           #temp_text2 := #Cfg_MessagePrefix.MessagePrefix[#temp_Language];
           IF LEN(#temp_text2) = 0 THEN #temp_text2 := ' ';  END_IF;

           #temp_text3 := #Cfg_Event.Message[#temp_Language];
           IF LEN(#temp_text3) = 0 THEN #temp_text3 := ' ';  END_IF;

        #In_EventStatus.Sts_Events[#Event_Number].Message := CONCAT(IN1 := #temp_text1, IN2 := #temp_text2, IN3 := #temp_text3);   // CONCAT (Cfg_MessagePrefix, Cfg_Event.Message);    
        //  #In_EventStatus.Sts_Events[#Event_Number].Message := CONCAT(IN1 := #temp_text1, IN2 := #Cfg_MessagePrefix.Language[#temp_Language], IN3 := #Cfg_Event.Message[#temp_Language]);   // CONCAT (Cfg_MessagePrefix, Cfg_Event.Message); 

           #In_EventStatus.Sts_Events[#Event_Number].Trigger := TRUE;                      // Set trigger to 1 
           #In_EventStatus.Sts_Events[#Event_Number].DateTime := #Event_CurDateTime;         // Update with the current time
           #In_EventStatus.Sts_Events[#Event_Number].AckDateTime := DT#1990-1-1-0:0:0.0;       // clear the acknowledge time value 
           END_IF;

      #Sts_Active   := TRUE;                            // set the status active bit
      #Sts_Latched  := TRUE;                            // set the status latched bit
      #In_EventStatus.Wrk_UpdateEventListID := #In_EventStatus.Wrk_UpdateEventListID+1;  // increment the work update listID


       CASE DINT_TO_INT(#Cfg_Event.Category) OF                     // set the appropriate category lateched bit 
           0: #In_EventStatus.Sts_Category_0_Latched :=1;
           1: #In_EventStatus.Sts_Category_1_Latched :=1;
           2: #In_EventStatus.Sts_Category_2_Latched :=1;
           3: #In_EventStatus.Sts_Category_3_Latched :=1;
           4: #In_EventStatus.Sts_Category_4_Latched :=1;
           5: #In_EventStatus.Sts_Category_5_Latched :=1;
           6: #In_EventStatus.Sts_Category_6_Latched :=1;
           7: #In_EventStatus.Sts_Category_7_Latched :=1;
           8: #In_EventStatus.Sts_Category_8_Latched :=1;
           9: #In_EventStatus.Sts_Category_9_Latched :=1;
       END_CASE;
   END_IF;                            // End "IF NOT (Sts_Active)"


   END_IF;                             // End "IF NOT(EnableIn) "


   //----------------------------------------------------- 
   ENO:= true;          // Set the ENO output
END_FUNCTION_BLOCK

FUNCTION_BLOCK "FB_TR88_CPG_EventManager"   // FB3102, SCL
TITLE = PackML EventManager (TR88 CPG Template)
{ S7_Optimized_Access := 'TRUE' }
AUTHOR : FoodBev
FAMILY : ISATR88e
NAME : EventMgr
VERSION : 1.81
// Takes the event information from the control modules (from FB_Event) and will create one list of events for the equipment module. It summarizes the data by finding the equipment module first out event and summarizes which category of events are active. This FB will also send reset commands to unlatch the control module events. Only one instance of this FB should be programmed per equipment module for each event type, for example one for alarms, one for warnings, etc.
   VAR_INPUT
      Cmd_Reset : Bool;   // Reset Command
      Cmd_ClearFirstOutEvents : Bool;   // Command to clear First Out events
      FirstScanBit : Bool;   // Bit used to tell logic that this is the firt scan of PLC
      Cfg_MessagePrefix : "UDT_TR88_CPG_Message_Prefix";   // Message Prefix value for event messages multi-lingual
      Cfg_Language : Int;   // Current Langage: 0=EN, 1=SP/ES, 2=DE, 3=FR, 4=IT
   END_VAR
   VAR_OUTPUT
      Sts_Category_0_Latched : Bool;   // Event Category Status (on until reset cmd) - CAT 0
      Sts_Category_1_Latched : Bool;   // Event Category Status (on until reset cmd) - CAT 1
      Sts_Category_2_Latched : Bool;   // Event Category Status (on until reset cmd) - CAT 2
      Sts_Category_3_Latched : Bool;   // Event Category Status (on until reset cmd) - CAT 3
      Sts_Category_4_Latched : Bool;   // Event Category Status (on until reset cmd) - CAT 4
      Sts_Category_5_Latched : Bool;   // Event Category Status (on until reset cmd) - CAT 5
      Sts_Category_6_Latched : Bool;   // Event Category Status (on until reset cmd) - CAT 6
      Sts_Category_7_Latched : Bool;   // Event Category Status (on until reset cmd) - CAT 7
      Sts_Category_8_Latched : Bool;   // Event Category Status (on until reset cmd) - CAT 8
      Sts_Category_9_Latched : Bool;   // Event Category Status (on until reset cmd) - CAT 9
      Sts_Category_0_NotLatched : Bool;   // Event Cat Status, not latched (=active event status) - CAT 0
      Sts_Category_1_NotLatched : Bool;   // Event Cat Status, not latched (=active event status) - CAT 1
      Sts_Category_2_NotLatched : Bool;   // Event Cat Status, not latched (=active event status) - CAT 2
      Sts_Category_3_NotLatched : Bool;   // Event Cat Status, not latched (=active event status) - CAT 3
      Sts_Category_4_NotLatched : Bool;   // Event Cat Status, not latched (=active event status) - CAT 4
      Sts_Category_5_NotLatched : Bool;   // Event Cat Status, not latched (=active event status) - CAT 5
      Sts_Category_6_NotLatched : Bool;   // Event Cat Status, not latched (=active event status) - CAT 6
      Sts_Category_7_NotLatched : Bool;   // Event Cat Status, not latched (=active event status) - CAT 7
      Sts_Category_8_NotLatched : Bool;   // Event Cat Status, not latched (=active event status) - CAT 8
      Sts_Category_9_NotLatched : Bool;   // Event Cat Status, not latched (=active event status) - CAT 9
      Sts_NumEvents : Int;   // Number of event in the In_EventStatus list
      Sts_CurrentActiveEvent : Bool;   // Status - TRUE = if any active events
      Sts_error : Bool;   // FB Error exist
      Sts_errorCode : DInt;   // FB Error code
   END_VAR
   VAR_IN_OUT
      In_EventStatus : "UDT_TR88_CPG_EventStatus";   // Working event list data section
   END_VAR
   VAR
      EventCategory : Int;
      Index_AllEvents : Int;
      Index_ClearActiveEvents : Int;
      Index_ClearFirstOut : Int;
      NumEvents : Int;   // Max # of Events
      Prev_CmdReset : Bool;
      Prev_NumEvents : Int;
      Prev_UpdateEventListID : Int;
      UpdateEventList : Bool;
      ZeroEvent : "UDT_TR88_CPG_Event";   // Null Event
   END_VAR
   VAR_TEMP
      "step" : Int;
      temp_text1 : String[30];
      temp_text2 : String[30];
      tempAnyPointer : DInt;   // temp Any poninter for FC_Array_Length call.
   END_VAR
BEGIN
   // ============================================================================ 
   // FUNCTION_BLOCK "FB_PMLe_EventManager"  
   // ---------------------------------------------------------------------------
   // Siemens Industry, Inc.
   // Food & Beverage VSS
   // ---------------------------------------------------------------------------
   // FUNCTIONALITY:  
   // Function Block to control EventManager function.
   // ---------------------------------------------------------------------------
   // change log table:
   // version        date          expert in charge        changes applied
   //  1.7         2012-08-22          M.Pieper           Matches Rev 1.7
   //                                                     Added Multi-Lingual support
   //  1.8       2013.07.31            M.Pieper           Removed EM message prefix logic
   //  1.81      2015-01-27            M.Pieper           Updated S7-1500 Array Size Logic.
   // ===========================================================================
   (*
   THIS SOFTWARE IS PROVIDED "AS IS" AND WITHOUT WARRANTIES OF ANY KIND, WHETHER EXPRESS OR IMPLIED.

   General information -
       Note :  the standard applications are NOT binding AND DO NOT claim TO be complete regarding configuration, equipment OR any eventuality which may arise. 
       The standard applications DO NOT represent specific customer solutions, but are only intended TO provide support FOR typical tasks. You are responsible 
       FOR the proper operation OF the described products. These standard applications DO NOT relieve you OF your responsibility regarding the safe handling 
       when using, installing operating AND maintaining the equipment. BY using these standard applications, you agree that Siemens cannot be made liable FOR 
       possible damage beyond the mentioned liability clause. We reserve the right TO make changes AND revisions TO these standard applications at Any Time 
       without prior notice. In the CASE OF Any differences between the suggestions made in these standard applications AND other publications from Siemens, 
       such as catalogs, the contents OF the other documentation have priority.

   Warranty conditions, liability, AND support -
      IF the application has been made available free OF charge, the following applies:
      * We DO NOT provide a warranty FOR Any OF the information contained in this document.
      * All other rights AND claims against Siemens AG irrespective OF legal basis are excluded. In particular claims FOR damages against Siemens AG 
      in the CASE OF Product outage, downtime, loss OF profit, either directly, indirectly OR consequential damage are excluded.
      * This does NOT apply when liability is compulsory BY law, e. g. in the CASE OF the Product liability act, premeditation, an act OF gross negligence 
      BY superiors AND managerial staff OF Siemens AG OR in cases OF fraudulent concealment OF defects.
      * This limitation OF liability also applies TO sub-contractors, suppliers, delegates, superiors AND managerial staff OF Siemens AG.
      German law shall apply TO this agreement FOR customers with head offices in Germany; Swiss law FOR customers with head offices outside Germany. 
      Application OF the United Nations Convention on Contracts FOR the International Sale OF Goods as OF 11.04.1980 (CISG) is excluded.
   *)

   // ===========================================================================
   //  Begin the LOGIC section:
   // First Scan Logic Logic (only ran on 1st scan of PLC)
   IF #FirstScanBit THEN                   //  First Scan bit set?
       #In_EventStatus.Wrk_ResetID := #In_EventStatus.Wrk_ResetID + 1;            // increment the Work Reset ID
       #In_EventStatus.Wrk_UpdateEventListID := #In_EventStatus.Wrk_UpdateEventListID + 1; // increment the Work UpdateList ID
       #In_EventStatus.Sts_NumAllEvents := 0;                                        // Reset the number of all events value
       // Determine the Number of Sts_Events for given alarm/warning area
       // S7-1500 Code: 
       "FC_ArrayLength_S7-1500"(Array_ToBe_Sized := #In_EventStatus.Sts_Events,
                                ArraySize => #In_EventStatus.Wrk_EventArraySize);
       RETURN;                            // Exit the FB call
   END_IF;                              // End the first scan section


   //---------------------------------------------------------------------------------
   // Main Logic Section

   // Update the message prefix for the current language
   #In_EventStatus.Wrk_LanguageSelection := #Cfg_Language;
   #In_EventStatus.Wrk_MessagePrefix := #Cfg_MessagePrefix.MessagePrefix[#In_EventStatus.Wrk_LanguageSelection];

   // Upon a reset command, reset the latched status bits and clear the event list
   IF #Cmd_Reset THEN
       #In_EventStatus.Sts_Category_0_Latched := 0;
       #In_EventStatus.Sts_Category_1_Latched := 0;
       #In_EventStatus.Sts_Category_2_Latched := 0;
       #In_EventStatus.Sts_Category_3_Latched := 0;
       #In_EventStatus.Sts_Category_4_Latched := 0;
       #In_EventStatus.Sts_Category_5_Latched := 0;
       #In_EventStatus.Sts_Category_6_Latched := 0;
       #In_EventStatus.Sts_Category_7_Latched := 0;
       #In_EventStatus.Sts_Category_8_Latched := 0;
       #In_EventStatus.Sts_Category_9_Latched := 0;

       IF NOT (#Prev_CmdReset) THEN                             // Clear the zero event
           #In_EventStatus.Out_ZeroEvent := #ZeroEvent;
           // String seperation variable not added.
       END_IF;
   END_IF;                      // End IF Cmd_Reset.... 


   // Clear first out events - for alarms, this is typically done once the machine starts    
   IF #Cmd_ClearFirstOutEvents AND NOT (#Sts_CurrentActiveEvent) THEN
       #In_EventStatus.Sts_FirstOutEvent := #In_EventStatus.Out_ZeroEvent;
       FOR #Index_ClearFirstOut := 0 TO 9 BY 1 DO
           #In_EventStatus.Sts_FirstOutEventCat[#Index_ClearFirstOut] := #In_EventStatus.Out_ZeroEvent;
       END_FOR;
   END_IF;

   // Determine the maximum number of event that can be stored in the array.  It is assumed that the input array
   // size is equal to the output array size!!
   IF (#Cmd_Reset AND (NOT #Prev_CmdReset)) OR (#In_EventStatus.Wrk_EventArraySize = 0) THEN
       // Determine the Number of Sts_Events for given alarm/warning area
       // S7-300 Code:
       // UDT_Event = 66 bytes in length
       // #tempAnyPointer := #In_EventStatus.Sts_Events;    // temp Any Pointer for FC_ArrrayLength call.
       // "FC_ArrayLength"(ArraySource:=#tempAnyPointer, ArrayLength:=66, SIZE=> #In_EventStatus.Wrk_EventArraySize);
       // 
       // S7-1500 Code: (TEST)
       //   VariantPut(SRC := #In_EventStatus.Sts_Events,
       //              DST := #temp_varArrayLengthPntr);              // Link input array to variant datatype.

       //              IF IS_ARRAY(#temp_varArrayLengthPntr) THEN                // Determine the length of the array...
       //                  #In_EventStatus.Wrk_EventArraySize := CountOfElements(#temp_varArrayLengthPntr);
       //              END_IF;
       // S7-1500 Code: 
       "FC_ArrayLength_S7-1500"(Array_ToBe_Sized := #In_EventStatus.Sts_Events,
                                ArraySize => #In_EventStatus.Wrk_EventArraySize);
   END_IF;

   //Determine if the event list needs updating    
   IF #In_EventStatus.Wrk_UpdateEventListID <> #Prev_UpdateEventListID THEN
       #Prev_UpdateEventListID := #In_EventStatus.Wrk_UpdateEventListID;
       #UpdateEventList := true;
   END_IF;

   IF #UpdateEventList THEN
       #UpdateEventList := false;
       // Update Event outputs and status
       // First clear the not lateched staus bits and total number of events.
       // This instruction will find the events in the coming rungs
       #Sts_errorCode := 0;
       #Sts_NumEvents := #In_EventStatus.Sts_NumAllEvents;
       #Sts_CurrentActiveEvent := false;
       #Sts_Category_0_NotLatched := false;
       #Sts_Category_1_NotLatched := false;
       #Sts_Category_2_NotLatched := false;
       #Sts_Category_3_NotLatched := false;
       #Sts_Category_4_NotLatched := false;
       #Sts_Category_5_NotLatched := false;
       #Sts_Category_6_NotLatched := false;
       #Sts_Category_7_NotLatched := false;
       #Sts_Category_8_NotLatched := false;
       #Sts_Category_9_NotLatched := false;

       //Determine if the number of events is greater than the max array size        
       //if so, then report error
       #NumEvents := #In_EventStatus.Sts_NumAllEvents;         // xxx
       IF #NumEvents > #In_EventStatus.Wrk_EventArraySize THEN
           #NumEvents := #In_EventStatus.Wrk_EventArraySize;  // 
           IF (#Sts_errorCode = 0) THEN                   // Update status error code
               #Sts_errorCode := 1;
           END_IF;
       END_IF;
       #In_EventStatus.Sts_NumEvents := #NumEvents;

       //Go Through the event array to cpature first fault event and perform STRING management        
       #Index_AllEvents := 0;
       FOR #Index_AllEvents := 0 TO #NumEvents - 1 DO
           // Check to see if any event is currently still active
           IF (#In_EventStatus.Sts_Events[#Index_AllEvents].Trigger) THEN   // 
               #Sts_CurrentActiveEvent := true;
           END_IF;

           //Store event category for logic later in code
           // EventCategory := In_EventStatus.Sts_Events[Index_allEvents].Category;  //From V1.2
           IF (#In_EventStatus.Sts_Events[#Index_AllEvents].Category >= 0) AND (#In_EventStatus.Sts_Events[#Index_AllEvents].Category <= 9) THEN
               #EventCategory := #In_EventStatus.Sts_Events[#Index_AllEvents].Category;
           ELSE
               #EventCategory := 0;
               IF (#Sts_errorCode = 0) THEN                   // Update status error code
                   #Sts_errorCode := 2;
               END_IF;         // end "IF (Sts_ErrorCode=0)"
           END_IF;             // end "IF (In_EventStatus.Sts_Events[Inde..."    

           // Set the First Out Event
           IF NOT (#In_EventStatus.Sts_FirstOutEvent.Trigger) THEN
               #In_EventStatus.Sts_FirstOutEvent := #In_EventStatus.Sts_Events[#Index_AllEvents];
               #In_EventStatus.Sts_FirstOutEvent.Trigger := True;
               // Clean up the ASCII characte strings - not needed
           END_IF;

           // Set the First Out Events by category
           IF NOT (#In_EventStatus.Sts_FirstOutEventCat[#EventCategory].Trigger) THEN
               #In_EventStatus.Sts_FirstOutEventCat[#EventCategory] := #In_EventStatus.Sts_Events[#Index_AllEvents];
               #In_EventStatus.Sts_FirstOutEventCat[#EventCategory].Trigger := True;
               // Clean up the ASCII characte strings - not needed
           END_IF;

           // Add message prefix to active event arrays


           //Category Event Status            
           CASE DINT_TO_INT(#In_EventStatus.Sts_Events[#Index_AllEvents].Category) OF
               0:  #Sts_Category_0_NotLatched := #In_EventStatus.Sts_Events[#Index_AllEvents].Trigger;
               1:  #Sts_Category_1_NotLatched := (#Sts_Category_1_NotLatched OR #In_EventStatus.Sts_Events[#Index_AllEvents].Trigger);
               2:  #Sts_Category_2_NotLatched := (#Sts_Category_2_NotLatched OR #In_EventStatus.Sts_Events[#Index_AllEvents].Trigger);
               3:  #Sts_Category_3_NotLatched := (#Sts_Category_3_NotLatched OR #In_EventStatus.Sts_Events[#Index_AllEvents].Trigger);
               4:  #Sts_Category_4_NotLatched := (#Sts_Category_4_NotLatched OR #In_EventStatus.Sts_Events[#Index_AllEvents].Trigger);
               5:  #Sts_Category_5_NotLatched := (#Sts_Category_5_NotLatched OR #In_EventStatus.Sts_Events[#Index_AllEvents].Trigger);
               6:  #Sts_Category_6_NotLatched := (#Sts_Category_6_NotLatched OR #In_EventStatus.Sts_Events[#Index_AllEvents].Trigger);
               7:  #Sts_Category_7_NotLatched := (#Sts_Category_7_NotLatched OR #In_EventStatus.Sts_Events[#Index_AllEvents].Trigger);
               8:  #Sts_Category_8_NotLatched := (#Sts_Category_8_NotLatched OR #In_EventStatus.Sts_Events[#Index_AllEvents].Trigger);
               9:  #Sts_Category_9_NotLatched := (#Sts_Category_9_NotLatched OR #In_EventStatus.Sts_Events[#Index_AllEvents].Trigger);
           END_CASE;  // End of DINT_TO_INT(In_EventStatus.sts_events[Ind....


       END_FOR;

       // set the status bits
       #Sts_Category_0_Latched := #In_EventStatus.Sts_Category_0_Latched;
       #Sts_Category_1_Latched := #In_EventStatus.Sts_Category_1_Latched;
       #Sts_Category_2_Latched := #In_EventStatus.Sts_Category_2_Latched;
       #Sts_Category_3_Latched := #In_EventStatus.Sts_Category_3_Latched;
       #Sts_Category_4_Latched := #In_EventStatus.Sts_Category_4_Latched;
       #Sts_Category_5_Latched := #In_EventStatus.Sts_Category_5_Latched;
       #Sts_Category_6_Latched := #In_EventStatus.Sts_Category_6_Latched;
       #Sts_Category_7_Latched := #In_EventStatus.Sts_Category_7_Latched;
       #Sts_Category_8_Latched := #In_EventStatus.Sts_Category_8_Latched;
       #Sts_Category_9_Latched := #In_EventStatus.Sts_Category_9_Latched;

       #In_EventStatus.Sts_Category_0_NotLatched := #Sts_Category_0_NotLatched;
       #In_EventStatus.Sts_Category_1_NotLatched := #Sts_Category_1_NotLatched;
       #In_EventStatus.Sts_Category_2_NotLatched := #Sts_Category_2_NotLatched;
       #In_EventStatus.Sts_Category_3_NotLatched := #Sts_Category_3_NotLatched;
       #In_EventStatus.Sts_Category_4_NotLatched := #Sts_Category_4_NotLatched;
       #In_EventStatus.Sts_Category_5_NotLatched := #Sts_Category_5_NotLatched;
       #In_EventStatus.Sts_Category_6_NotLatched := #Sts_Category_6_NotLatched;
       #In_EventStatus.Sts_Category_7_NotLatched := #Sts_Category_7_NotLatched;
       #In_EventStatus.Sts_Category_8_NotLatched := #Sts_Category_8_NotLatched;
       #In_EventStatus.Sts_Category_9_NotLatched := #Sts_Category_9_NotLatched;

       #In_EventStatus.Sts_CurrentActiveEvent := #Sts_CurrentActiveEvent;
   END_IF;

   // Clear the remaining inactive bits    
   IF #Prev_NumEvents > #In_EventStatus.Sts_NumEvents THEN
       FOR #Index_ClearActiveEvents := #In_EventStatus.Sts_NumEvents TO #Prev_NumEvents - 1 DO
           #In_EventStatus.Sts_Events[#Index_ClearActiveEvents] := #In_EventStatus.Out_ZeroEvent;
       END_FOR;
   END_IF;

   // Clear the number of input events in the case where some control module events are not being actively scanned.    
   IF #Cmd_Reset AND ((#In_EventStatus.Sts_CurrentActiveEvent) OR (#In_EventStatus.Sts_NumEvents > 0) OR (NOT #Prev_CmdReset)) THEN
       #In_EventStatus.Wrk_ResetID := #In_EventStatus.Wrk_ResetID + 1;
       #In_EventStatus.Wrk_UpdateEventListID := #In_EventStatus.Wrk_UpdateEventListID + 1;
       #In_EventStatus.Sts_NumAllEvents := 0;
   END_IF;

   #Prev_NumEvents := #In_EventStatus.Sts_NumEvents;
   #Prev_CmdReset := #Cmd_Reset;
   #Sts_error := (#Sts_errorCode <> 0);

   //----------------------------------------------------- 
   ENO := true;   // Set the ENO output
END_FUNCTION_BLOCK

FUNCTION_BLOCK "FB_TR88_CPG_EventSumBegin"   // FB3103, SCL
TITLE = PackML Event Summation Begin (TR88 CPG Template)
{ S7_Optimized_Access := 'TRUE' }
AUTHOR : FoodBev
FAMILY : ISATR88e
NAME : EvSumBeg
VERSION : 1.2
// Summarizes the data from the equipment modules (from FB_EventManager) and will create one list of events for the unit machine. It summarizes the data by finding the unit machine first out event and summarizes which category of events are active. FB_EventSummationBegin initializes the summation, and FB_EventSummationEnd finalizes the summation.
   VAR_INPUT
      FirstScanBit : Bool;   // Bit used to tell logic that this is the firt scan of PLC
   END_VAR
   VAR_IN_OUT
      Sts_EventSummation : "UDT_TR88_CPG_EventSummation";   // Working event list data section
   END_VAR
   VAR
      Index : Int;   // temp value needed with FOR loop
      ZeroEvent : "UDT_TR88_CPG_Event";   // Null Event
   END_VAR
   VAR_TEMP
      tempAnyPointer : DInt;   // temp Any poninter for FC_Array_Length call.
      index_1 : Int;   // index counter
   END_VAR
BEGIN
   // ============================================================================ 
   // FUNCTION_BLOCK "FB_PMLe_EventSumBegin"  
   // ---------------------------------------------------------------------------
   // Siemens Industry, Inc.
   // Food & Beverage VSS
   // ---------------------------------------------------------------------------
   // FUNCTIONALITY:  
   // Summarizes the data from the equipment modules (from FB_EventManager) and will create one list of events for the unit machine.
   // It summarizes the data by finding the unit machine first out event and summarizes which category of events are active.
   // FB_EventSummationBegin initializes the summation, and FB_EventSummationEnd finalizes the summation.
   // ---------------------------------------------------------------------------
   // change log table:
   // version        date          expert in charge        changes applied
   // 
   //  1.1         2012-08-20        Mike Pieper        Matches Rev 1.1
   //  1.11        2015-01-27        Mike Pieper        Updated S7-1500 Array Size Logic.
   //  1.2         2015.04.01        Mike Pieper        TR88.00.02 Edition 2 Release. 
   // ===========================================================================
   (*
   THIS SOFTWARE IS PROVIDED "AS IS" AND WITHOUT WARRANTIES OF ANY KIND, WHETHER EXPRESS OR IMPLIED.

   General information -
       Note :  the standard applications are NOT binding AND DO NOT claim TO be complete regarding configuration, equipment OR any eventuality which may arise. 
       The standard applications DO NOT represent specific customer solutions, but are only intended TO provide support FOR typical tasks. You are responsible 
       FOR the proper operation OF the described products. These standard applications DO NOT relieve you OF your responsibility regarding the safe handling 
       when using, installing operating AND maintaining the equipment. BY using these standard applications, you agree that Siemens cannot be made liable FOR 
       possible damage beyond the mentioned liability clause. We reserve the right TO make changes AND revisions TO these standard applications at Any Time 
       without prior notice. In the CASE OF Any differences between the suggestions made in these standard applications AND other publications from Siemens, 
       such as catalogs, the contents OF the other documentation have priority.

   Warranty conditions, liability, AND support -
      IF the application has been made available free OF charge, the following applies:
      * We DO NOT provide a warranty FOR Any OF the information contained in this document.
      * All other rights AND claims against Siemens AG irrespective OF legal basis are excluded. In particular claims FOR damages against Siemens AG 
      in the CASE OF Product outage, downtime, loss OF profit, either directly, indirectly OR consequential damage are excluded.
      * This does NOT apply when liability is compulsory BY law, e. g. in the CASE OF the Product liability act, premeditation, an act OF gross negligence 
      BY superiors AND managerial staff OF Siemens AG OR in cases OF fraudulent concealment OF defects.
      * This limitation OF liability also applies TO sub-contractors, suppliers, delegates, superiors AND managerial staff OF Siemens AG.
      German law shall apply TO this agreement FOR customers with head offices in Germany; Swiss law FOR customers with head offices outside Germany. 
      Application OF the United Nations Convention on Contracts FOR the International Sale OF Goods as OF 11.04.1980 (CISG) is excluded.
   *)

   // ===========================================================================
   // Begin the Firt Scan / Initialize LOGIC section:
   IF #FirstScanBit THEN
       "FC_ArrayLength_S7-1500"(Array_ToBe_Sized := #Sts_EventSummation.Sts_Events,
                                ArraySize => #Sts_EventSummation.Wrk_EventArraySize);

       FOR #Index := 0 TO (#Sts_EventSummation.Wrk_EventArraySize-1) DO
           #Sts_EventSummation.Sts_Events[#Index] := #ZeroEvent;
       END_FOR;

   END_IF;
   // End of First Scan Section

   // Begin the LOGIC section:
   // Initialize the summation - This FB is to be called before the numerous "FB_PG_EventSum" calls.

   // Clear the first out event
   #Sts_EventSummation.Sts_FirstOutEvent := #ZeroEvent;

   // Clear the first out event category arrays  
   FOR #Index := 0 TO 9 DO
       #Sts_EventSummation.Sts_FirstOutEventCat[#Index] := #ZeroEvent;
   END_FOR;

   // UDT_Event = 66 bytes in length
   // Determine the Number of Sts_Events for given alarm/warning area
   // S7-300 Logic:
   // #tempAnyPointer := #Sts_EventSummation.Sts_Events;    // temp Any Pointer for FC_ArrrayLength call.
   // "FC_ArrayLength"(ArraySource:= #tempAnyPointer, ArrayLength:=66, SIZE=> #Sts_EventSummation.Wrk_EventArraySize);
   // S7-1500 Logic:
   "FC_ArrayLength_S7-1500"(Array_ToBe_Sized := #Sts_EventSummation.Sts_Events,
                            ArraySize => #Sts_EventSummation.Wrk_EventArraySize);
   // Clear the number of events
   #Sts_EventSummation.Sts_NumEvents := 0;            // set the number of events to 0.

   // Clear the output category status bits
   #Sts_EventSummation.Wrk_Category_0_Latched := FALSE;
   #Sts_EventSummation.Wrk_Category_1_Latched := FALSE;
   #Sts_EventSummation.Wrk_Category_2_Latched := FALSE;
   #Sts_EventSummation.Wrk_Category_3_Latched := FALSE;
   #Sts_EventSummation.Wrk_Category_4_Latched := FALSE;
   #Sts_EventSummation.Wrk_Category_5_Latched := FALSE;
   #Sts_EventSummation.Wrk_Category_6_Latched := FALSE;
   #Sts_EventSummation.Wrk_Category_7_Latched := FALSE;
   #Sts_EventSummation.Wrk_Category_8_Latched := FALSE;
   #Sts_EventSummation.Wrk_Category_9_Latched := FALSE;
   #Sts_EventSummation.Wrk_Category_0_NotLatched := FALSE;
   #Sts_EventSummation.Wrk_Category_1_NotLatched := FALSE;
   #Sts_EventSummation.Wrk_Category_2_NotLatched := FALSE;
   #Sts_EventSummation.Wrk_Category_3_NotLatched := FALSE;
   #Sts_EventSummation.Wrk_Category_4_NotLatched := FALSE;
   #Sts_EventSummation.Wrk_Category_5_NotLatched := FALSE;
   #Sts_EventSummation.Wrk_Category_6_NotLatched := FALSE;
   #Sts_EventSummation.Wrk_Category_7_NotLatched := FALSE;
   #Sts_EventSummation.Wrk_Category_8_NotLatched := FALSE;
   #Sts_EventSummation.Wrk_Category_9_NotLatched := FALSE;
   #Sts_EventSummation.Wrk_CurrentActiveEvent := FALSE;

   //  ------------------------------------------------------------------

   ENO := true;   // Set the ENO output
END_FUNCTION_BLOCK

FUNCTION_BLOCK "FB_TR88_CPG_EventSum"   // FB3104, SCL
TITLE = PackML Event Summation (TR88 CPG Template)
{ S7_Optimized_Access := 'TRUE' }
AUTHOR : FoodBev
FAMILY : ISATR88e
NAME : EventSum
VERSION : 2.00
// Summarizes the data from the equipment modules (from FB_EventManager) and will create one list of events for the unit machine. It summarizes the data by finding the unit machine first out event and summarizes which category of events are active. FB_EventSummationBegin initializes the summation, and FB_EventSummationEnd finalizes the summation.
   VAR_OUTPUT
      Sts_NumEvents : Int;   // Status - Number of active events
      Sts_Category_0_Latched : Bool;   // Status - Latched Event - Cat. 0
      Sts_Category_1_Latched : Bool;   // Status - Latched Event - Cat. 1
      Sts_Category_2_Latched : Bool;   // Status - Latched Event - Cat. 2
      Sts_Category_3_Latched : Bool;   // Status - Latched Event - Cat. 3
      Sts_Category_4_Latched : Bool;   // Status - Latched Event - Cat. 4
      Sts_Category_5_Latched : Bool;   // Status - Latched Event - Cat. 5
      Sts_Category_6_Latched : Bool;   // Status - Latched Event - Cat. 6
      Sts_Category_7_Latched : Bool;   // Status - Latched Event - Cat. 7
      Sts_Category_8_Latched : Bool;   // Status - Latched Event - Cat. 8
      Sts_Category_9_Latched : Bool;   // Status - Latched Event - Cat. 9
      Sts_Category_0_NotLatched : Bool;   // Status - NotLatched (Active) Event - Cat. 0
      Sts_Category_1_NotLatched : Bool;   // Status - NotLatched (Active) Event - Cat. 1
      Sts_Category_2_NotLatched : Bool;   // Status - NotLatched (Active) Event - Cat. 2
      Sts_Category_3_NotLatched : Bool;   // Status - NotLatched (Active) Event - Cat. 3
      Sts_Category_4_NotLatched : Bool;   // Status - NotLatched (Active) Event - Cat. 4
      Sts_Category_5_NotLatched : Bool;   // Status - NotLatched (Active) Event - Cat. 5
      Sts_Category_6_NotLatched : Bool;   // Status - NotLatched (Active) Event - Cat. 6
      Sts_Category_7_NotLatched : Bool;   // Status - NotLatched (Active) Event - Cat. 7
      Sts_Category_8_NotLatched : Bool;   // Status - NotLatched (Active) Event - Cat. 8
      Sts_Category_9_NotLatched : Bool;   // Status - NotLatched (Active) Event - Cat. 9
      Sts_CurrentActiveEvent : Bool;   // Active Event Exists
      Sts_Error : Bool;   // Error in FB
      Sts_ErrorCode : DInt;   // Error Code
   END_VAR
   VAR_IN_OUT
      In_EventStatus : "UDT_TR88_CPG_EventStatus";   // UDT of EventStatus
      Sts_EventSummation : "UDT_TR88_CPG_EventSummation";   // UDT of EventSummation
   END_VAR
   VAR
      Cfg_MaxEvents : Int;   // number of events used from In_EventStatus array.
      Index : Int;
      NumEvents : Int;
      Prev_NumAllEvents : Int;
      UpdateEventList : Bool;
      WriteData : Bool;
      prev_updateEventListID : Int;
      error_RTC : Int;   // Error code for reading of Real Time Clock
      Event_CurDateTime : Date_And_Time;   // temp value for current date & time
      Compare1st_InNew : Bool;
      Compare1st_StsNew : Bool;
      Compare1stCat_InNew : Bool;
      Compare1stCat_StsNew : Bool;
   END_VAR
   VAR_TEMP
      temp_DT_1 : Date_And_Time;   // Temp Date & Time value
      temp_DT_2 : Date_And_Time;   // Temp Date & Time value
      tempAnyPointer : DInt;
   END_VAR
BEGIN
   // ============================================================================ 
   // FUNCTION_BLOCK "FB_PMLe_EventSum"  
   // ---------------------------------------------------------------------------
   // Siemens Industry, Inc.
   // Food & Beverage VSS
   // ---------------------------------------------------------------------------
   // FUNCTIONALITY:   
   // Summarizes the data from the equipment modules (from FB_EventManager) and will create one list of events for the unit machine.
   // It summarizes the data by finding the unit machine first out event and summarizes which category of events are active.
   // FB_EventSummationBegin initializes the summation, and FB_EventSummationEnd finalizes the summation.
   // ---------------------------------------------------------------------------
   // change log table:
   // version        date          expert in charge        changes applied
   //  1.5        2012-08-20        Mike Pieper        Matches Rev 1.5
   //  1.51       2015-01-27        Mike Pieper        Updated S7-1500 Array Size Logic.
   //  2.0        2015.04.01        Mike Pieper        TR88.00.02 Edition 2 Release.    
   // ===========================================================================
   (*
   THIS SOFTWARE IS PROVIDED "AS IS" AND WITHOUT WARRANTIES OF ANY KIND, WHETHER EXPRESS OR IMPLIED.

   General information -
       Note :  the standard applications are NOT binding AND DO NOT claim TO be complete regarding configuration, equipment OR any eventuality which may arise. 
       The standard applications DO NOT represent specific customer solutions, but are only intended TO provide support FOR typical tasks. You are responsible 
       FOR the proper operation OF the described products. These standard applications DO NOT relieve you OF your responsibility regarding the safe handling 
       when using, installing operating AND maintaining the equipment. BY using these standard applications, you agree that Siemens cannot be made liable FOR 
       possible damage beyond the mentioned liability clause. We reserve the right TO make changes AND revisions TO these standard applications at Any Time 
       without prior notice. In the CASE OF Any differences between the suggestions made in these standard applications AND other publications from Siemens, 
       such as catalogs, the contents OF the other documentation have priority.

   Warranty conditions, liability, AND support -
      IF the application has been made available free OF charge, the following applies:
      * We DO NOT provide a warranty FOR Any OF the information contained in this document.
      * All other rights AND claims against Siemens AG irrespective OF legal basis are excluded. In particular claims FOR damages against Siemens AG 
      in the CASE OF Product outage, downtime, loss OF profit, either directly, indirectly OR consequential damage are excluded.
      * This does NOT apply when liability is compulsory BY law, e. g. in the CASE OF the Product liability act, premeditation, an act OF gross negligence 
      BY superiors AND managerial staff OF Siemens AG OR in cases OF fraudulent concealment OF defects.
      * This limitation OF liability also applies TO sub-contractors, suppliers, delegates, superiors AND managerial staff OF Siemens AG.
      German law shall apply TO this agreement FOR customers with head offices in Germany; Swiss law FOR customers with head offices outside Germany. 
      Application OF the United Nations Convention on Contracts FOR the International Sale OF Goods as OF 11.04.1980 (CISG) is excluded.
   *)

   // ===========================================================================
   //  Begin the LOGIC section:

   #Sts_ErrorCode := 0;               // Set the status error code

   // Determine the Number of Sts_Events for given alarm/warning area
   // UDT_Event = 66 bytes in length
   // S7-300 Code:
   //#tempAnyPointer := #Sts_EventSummation.Sts_Events;    // temp Any Pointer for FC_ArrrayLength call.
   //"FC_ArrayLength"(ArraySource:= #tempAnyPointer, ArrayLength:=66, SIZE=> #Sts_EventSummation.Wrk_EventArraySize);
   //
   //#tempAnyPointer := #In_EventStatus.Sts_Events;    // temp Any Pointer for FC_ArrrayLength call.
   //"FC_ArrayLength"(ArraySource:= #tempAnyPointer, ArrayLength:=66, SIZE=> #Cfg_MaxEvents );  // the Number OF Sts_Events
   //
   // S7-1500 Code:
   "FC_ArrayLength_S7-1500"(Array_ToBe_Sized := #Sts_EventSummation.Sts_Events,
                            ArraySize => #Sts_EventSummation.Wrk_EventArraySize);
   // 
   "FC_ArrayLength_S7-1500"(Array_ToBe_Sized := #In_EventStatus.Sts_Events,
                            ArraySize => #Cfg_MaxEvents);

   #WriteData       :=0;               // set write data to false

   // Set First Out Event
   #temp_DT_1:=#In_EventStatus.Sts_FirstOutEvent.DateTime;                  // Date & Time of Sts_FirstOutEventCat[index].TimeEvent...
   IF #temp_DT_1 <> DT#1990-1-1-0:0:0.0 THEN                                // is In_EventStatus.Sts_FirstOutEvent.TimeEvent <> 0?
      #temp_DT_2:=#Sts_EventSummation.Sts_FirstOutEvent.DateTime;           // load the current value of the Sts_Eve..
         #WriteData:=0;                                                     // Reset the write data command.
         IF #temp_DT_2 = DT#1990-1-1-0:0:0.0 THEN                           // is Sts_EventSummation.Sts_FirstOutEvent.TimeEvent = 0? 
              #WriteData:=1;
         ELSIF #temp_DT_1 < #temp_DT_2 THEN                                  // is IN_event newer than Sts_event ?
              #WriteData:=1;
         END_IF;     // End "IF (EQ_DT(DT1:=Sts_"
   END_IF;         // End "IF (NOT(EQ_DT(DT1:=In_Ev"

   IF #WriteData THEN 
      #Sts_EventSummation.Sts_FirstOutEvent:=#In_EventStatus.Sts_FirstOutEvent;  // Update the First Fault event 
   END_IF; 

   // Set First Out Event by Category
   FOR #Index:= 0 TO 9 DO
       #temp_DT_1:=#In_EventStatus.Sts_FirstOutEventCat[#Index].DateTime;        // Date & Time of Sts_FirstOutEventCat[index].TimeEvent...
       IF #temp_DT_1 <> DT#1990-1-1-0:0:0.0 THEN                                // is In_EventStatus.Sts_FirstOutEvent.TimeEvent <> 0?
           #temp_DT_2:=#Sts_EventSummation.Sts_FirstOutEventCat[#Index].DateTime;          // load the current value of the Sts_Eve..
           #WriteData:=0;                   // Reset the write data command.
           IF #temp_DT_2 = DT#1990-1-1-0:0:0.0 THEN                              // is Sts_EventSummation.Sts_FirstOutEvent.TimeEvent = 0? 
               #WriteData:=1;
           ELSIF #temp_DT_1 < #temp_DT_2 THEN                                    // is IN_event newer than Sts_event ?
               #WriteData:=1;
           END_IF;     // End "IF (EQ_DT(DT1:=Sts_"
       END_IF;         // End "IF (NOT(EQ_DT(DT1:=In_Ev"

       IF #WriteData THEN 
           #Sts_EventSummation.Sts_FirstOutEventCat[#Index]:=#In_EventStatus.Sts_FirstOutEventCat[#Index];  // Update the First Fault event 
       END_IF; 
   END_FOR;     

   // ---------------------------------------------------------------
   // Set Active Events
   IF #In_EventStatus.Sts_NumEvents > 0 THEN 
           #NumEvents:=#In_EventStatus.Sts_NumEvents;
         IF (#Cfg_MaxEvents > 0) AND (#NumEvents>#Cfg_MaxEvents) THEN
               #NumEvents:=#Cfg_MaxEvents;
         END_IF;

         IF #NumEvents > (#Sts_EventSummation.Wrk_EventArraySize - #Sts_EventSummation.Sts_NumEvents) THEN
               #NumEvents:=#Sts_EventSummation.Wrk_EventArraySize-#Sts_EventSummation.Sts_NumEvents;
             IF (#Sts_ErrorCode=0)   THEN 
                   #Sts_ErrorCode:=1;
             END_IF;
         END_IF;                

       IF #NumEvents > 0 THEN
           FOR #Index:= 0 TO DINT_TO_INT(#NumEvents-1) DO  // 
               #Sts_EventSummation.Sts_Events[#Index+#Sts_EventSummation.Sts_NumEvents]:= #In_EventStatus.Sts_Events[#Index];
           END_FOR;
           #Sts_EventSummation.Sts_NumEvents:= #Sts_EventSummation.Sts_NumEvents + #NumEvents;
       END_IF;    
   END_IF;

   #Sts_NumEvents:=#Sts_EventSummation.Sts_NumEvents;

   // Set Category Bits
   #Sts_EventSummation.Wrk_Category_0_Latched := (#Sts_EventSummation.Wrk_Category_0_Latched OR #In_EventStatus.Sts_Category_0_Latched);
   #Sts_EventSummation.Wrk_Category_1_Latched := (#Sts_EventSummation.Wrk_Category_1_Latched OR #In_EventStatus.Sts_Category_1_Latched);
   #Sts_EventSummation.Wrk_Category_2_Latched := (#Sts_EventSummation.Wrk_Category_2_Latched OR #In_EventStatus.Sts_Category_2_Latched);
   #Sts_EventSummation.Wrk_Category_3_Latched := (#Sts_EventSummation.Wrk_Category_3_Latched OR #In_EventStatus.Sts_Category_3_Latched);
   #Sts_EventSummation.Wrk_Category_4_Latched := (#Sts_EventSummation.Wrk_Category_4_Latched OR #In_EventStatus.Sts_Category_4_Latched);
   #Sts_EventSummation.Wrk_Category_5_Latched := (#Sts_EventSummation.Wrk_Category_5_Latched OR #In_EventStatus.Sts_Category_5_Latched);
   #Sts_EventSummation.Wrk_Category_6_Latched := (#Sts_EventSummation.Wrk_Category_6_Latched OR #In_EventStatus.Sts_Category_6_Latched);
   #Sts_EventSummation.Wrk_Category_7_Latched := (#Sts_EventSummation.Wrk_Category_7_Latched OR #In_EventStatus.Sts_Category_7_Latched);
   #Sts_EventSummation.Wrk_Category_8_Latched := (#Sts_EventSummation.Wrk_Category_8_Latched OR #In_EventStatus.Sts_Category_8_Latched);
   #Sts_EventSummation.Wrk_Category_9_Latched := (#Sts_EventSummation.Wrk_Category_9_Latched OR #In_EventStatus.Sts_Category_9_Latched);

   #Sts_Category_0_Latched := #In_EventStatus.Sts_Category_0_Latched;
   #Sts_Category_1_Latched := #In_EventStatus.Sts_Category_1_Latched;
   #Sts_Category_2_Latched := #In_EventStatus.Sts_Category_2_Latched;
   #Sts_Category_3_Latched := #In_EventStatus.Sts_Category_3_Latched;
   #Sts_Category_4_Latched := #In_EventStatus.Sts_Category_4_Latched;
   #Sts_Category_5_Latched := #In_EventStatus.Sts_Category_5_Latched;
   #Sts_Category_6_Latched := #In_EventStatus.Sts_Category_6_Latched;
   #Sts_Category_7_Latched := #In_EventStatus.Sts_Category_7_Latched;
   #Sts_Category_8_Latched := #In_EventStatus.Sts_Category_8_Latched;
   #Sts_Category_9_Latched := #In_EventStatus.Sts_Category_9_Latched;

   #Sts_EventSummation.Wrk_Category_0_NotLatched := #Sts_EventSummation.Wrk_Category_0_NotLatched OR #In_EventStatus.Sts_Category_0_NotLatched;
   #Sts_EventSummation.Wrk_Category_1_NotLatched := #Sts_EventSummation.Wrk_Category_1_NotLatched OR #In_EventStatus.Sts_Category_1_NotLatched;
   #Sts_EventSummation.Wrk_Category_2_NotLatched := #Sts_EventSummation.Wrk_Category_2_NotLatched OR #In_EventStatus.Sts_Category_2_NotLatched;
   #Sts_EventSummation.Wrk_Category_3_NotLatched := #Sts_EventSummation.Wrk_Category_3_NotLatched OR #In_EventStatus.Sts_Category_3_NotLatched;
   #Sts_EventSummation.Wrk_Category_4_NotLatched := #Sts_EventSummation.Wrk_Category_4_NotLatched OR #In_EventStatus.Sts_Category_4_NotLatched;
   #Sts_EventSummation.Wrk_Category_5_NotLatched := #Sts_EventSummation.Wrk_Category_5_NotLatched OR #In_EventStatus.Sts_Category_5_NotLatched;
   #Sts_EventSummation.Wrk_Category_6_NotLatched := #Sts_EventSummation.Wrk_Category_6_NotLatched OR #In_EventStatus.Sts_Category_6_NotLatched;
   #Sts_EventSummation.Wrk_Category_7_NotLatched := #Sts_EventSummation.Wrk_Category_7_NotLatched OR #In_EventStatus.Sts_Category_7_NotLatched;
   #Sts_EventSummation.Wrk_Category_8_NotLatched := #Sts_EventSummation.Wrk_Category_8_NotLatched OR #In_EventStatus.Sts_Category_8_NotLatched;
   #Sts_EventSummation.Wrk_Category_9_NotLatched := #Sts_EventSummation.Wrk_Category_9_NotLatched OR #In_EventStatus.Sts_Category_9_NotLatched;

   #Sts_Category_0_NotLatched := #In_EventStatus.Sts_Category_0_NotLatched;
   #Sts_Category_1_NotLatched := #In_EventStatus.Sts_Category_1_NotLatched;
   #Sts_Category_2_NotLatched := #In_EventStatus.Sts_Category_2_NotLatched;
   #Sts_Category_3_NotLatched := #In_EventStatus.Sts_Category_3_NotLatched;
   #Sts_Category_4_NotLatched := #In_EventStatus.Sts_Category_4_NotLatched;
   #Sts_Category_5_NotLatched := #In_EventStatus.Sts_Category_5_NotLatched;
   #Sts_Category_6_NotLatched := #In_EventStatus.Sts_Category_6_NotLatched;
   #Sts_Category_7_NotLatched := #In_EventStatus.Sts_Category_7_NotLatched;
   #Sts_Category_8_NotLatched := #In_EventStatus.Sts_Category_8_NotLatched;
   #Sts_Category_9_NotLatched := #In_EventStatus.Sts_Category_9_NotLatched;

   #Sts_EventSummation.Wrk_CurrentActiveEvent := #Sts_EventSummation.Wrk_CurrentActiveEvent OR #In_EventStatus.Sts_CurrentActiveEvent;

   #Sts_CurrentActiveEvent := #In_EventStatus.Sts_CurrentActiveEvent;

   // Set Error Bit
   #Sts_Error:=(#Sts_ErrorCode<>0);

   //  ------------------------------------------------------------------
   ENO:= true;   // Set the ENO output
END_FUNCTION_BLOCK

FUNCTION_BLOCK "FB_TR88_CPG_EventSumEnd"   // FB3105, SCL
TITLE = PackML Event Summation End (TR88 CPG Template)
{ S7_Optimized_Access := 'TRUE' }
AUTHOR : FoodBev
FAMILY : ISATR88e
NAME : EvSumEnd
VERSION : 1.11
// Summarizes the data from the equipment modules (from FB_EventManager) and will create one list of events for the unit machine. It summarizes the data by finding the unit machine first out event and summarizes which category of events are active. FB_EventSummationBegin initializes the summation, and FB_EventSummationEnd finalizes the summation.
   VAR_IN_OUT
      Sts_EventSummation : "UDT_TR88_CPG_EventSummation";   // Working event list data section
   END_VAR
   VAR
      Index : Int;
      Prev_NumAllEvents : Int;   // temp value needed with FOR loop
      ZeroEvent : "UDT_TR88_CPG_Event";   // Null Event
   END_VAR
   VAR_TEMP
      ZeroEvent1 : "UDT_TR88_CPG_Event";   // null instance of UDT Event
      tempAnyPointer : DInt;
   END_VAR
BEGIN
   // ============================================================================ 
   // FUNCTION_BLOCK "FB_PMLe_EventSumEnd"    
   // ---------------------------------------------------------------------------
   // Siemens Industry, Inc.
   // Food & Beverage VMM
   // ---------------------------------------------------------------------------
   // FUNCTIONALITY:  
   // Summarizes the data from the equipment modules (from FB_EventManager) and will create one list of events for the unit machine.
   // It summarizes the data by finding the unit machine first out event and summarizes which category of events are active.
   // FB_EventSummationBegin initializes the summation, and FB_EventSummationEnd finalizes the summation.
   // ---------------------------------------------------------------------------
   // change log table:
   // version        date          expert in charge        changes applied
   // 
   //  1.1         2012-08-20          M.Pieper            Matches Rev 1.1
   //  1.11        2015-01-27          M.Pieper            Updated S7-1500 Array Size Logic. 
   // ===========================================================================
   (*
   THIS SOFTWARE IS PROVIDED "AS IS" AND WITHOUT WARRANTIES OF ANY KIND, WHETHER EXPRESS OR IMPLIED.

   General information -
       Note :  the standard applications are NOT binding AND DO NOT claim TO be complete regarding configuration, equipment OR any eventuality which may arise. 
       The standard applications DO NOT represent specific customer solutions, but are only intended TO provide support FOR typical tasks. You are responsible 
       FOR the proper operation OF the described products. These standard applications DO NOT relieve you OF your responsibility regarding the safe handling 
       when using, installing operating AND maintaining the equipment. BY using these standard applications, you agree that Siemens cannot be made liable FOR 
       possible damage beyond the mentioned liability clause. We reserve the right TO make changes AND revisions TO these standard applications at Any Time 
       without prior notice. In the CASE OF Any differences between the suggestions made in these standard applications AND other publications from Siemens, 
       such as catalogs, the contents OF the other documentation have priority.